// TIA Portal project "ljussennsor skåp" (V18)

(* hardware
DEVICE "S7-1200 station_1"  S7-1200 Station
   slot 0: "Rack_0"  S7-1200 Rack  Rack  V1.0
   slot 1: "PLC_1"  CPU 1212C DC/DC/DC  6ES7 212-1AE40-0XB0  V4.5
DEVICE "HMI_1"  TP900 Comfort
   slot 0: "HMI_1"  TP900 Comfort  6AV2 124-0JC01-0AX0  17.0.0.0
   slot 1: "HMI_RT_1"  TP900 Comfort  6AV2 124-0JC01-0AX0  17.0.0.0
   slot 5: "HMI_1.IE_CP_1"  PROFINET Interface  17.0.0.0
      slot 1: "PROFINET Interface_1"  PROFINET Interface
         slot 1: "Port_1"  Port
         slot 2: "Port_2"  Port
   slot 7: "HMI_1.MPI/DP_CP_1"  MPI/DP Interface  17.0.0.0
*)

// ===== PLC "PLC_1"  CPU 1212C DC/DC/DC =====

VAR_GLOBAL   // PLC tag table "Default tag table"
   "Tag_1" AT %I0.4 : Bool;
   "Tag_2" AT %I0.5 : Bool;
   "Tag_3" AT %I0.6 : Bool;
   "ok" AT %M0.7 : Bool;
END_VAR

VAR_GLOBAL   // PLC tag table "Analog_Tag"
   "Star/Button" AT %I0.0 : Bool;
   "Stop/Button" AT %I0.1 : Bool;
   "Reset/Button" AT %I0.2 : Bool;
   "light sensor" AT %IW64 : Int;
   "Green" AT %Q0.0 : Bool;   // Lamp
   "Red" AT %Q0.1 : Bool;   // Lamp
   "Yellow" AT %Q0.2 : Bool;   // Lamp
   "LEDLights" AT %Q0.3 : Bool;
END_VAR

DATA_BLOCK "data"   // DB1
{ S7_Optimized_Access := 'TRUE' }
VERSION : 0.1
   VAR
      normxstruct : Struct
         minval : Int := 0;
         maxval : Int := 27648;
         lightval : Int;
         normxoutput : Real;
      END_STRUCT;
      lightpercent : Struct
         percentofthelight : Real;
      END_STRUCT;
      calibratedvalues : Struct
         "2layermin" : Real;
         "2layermax" : Real;
      END_STRUCT;
      defaultvalues : Struct
         minimumvalue : Real := 87.9;
         maxvalue : Real := 86.2;
      END_STRUCT;
      startcalibration : Bool;
      finishedcalibration : Bool;
      hmibuttons : Struct
         hmistartbutton : Bool;
         hmiyellowbutton : Bool;
         hmiredbutton : Bool;
      END_STRUCT;
   END_VAR
BEGIN
END_DATA_BLOCK

// folder: System blocks/Program resources

DATA_BLOCK "IEC_Counter_0_DB_1"   // DB3
{ S7_Optimized_Access := 'TRUE' }
AUTHOR : Simatic
FAMILY : IEC
NAME : CNTR
VERSION : 1.0
// stored: InstanceOfName IEC_COUNTER
"IEC_COUNTER"
BEGIN
END_DATA_BLOCK

// folder: (top level)

FUNCTION "function" : Void   // FC1, LAD
{ S7_Optimized_Access := 'TRUE' }
VERSION : 0.1
   VAR_TEMP   // added for the SCL form of the ladder/FBD networks
      _w1 : Bool;
      _w2 : Bool;
      _w3 : Bool;
      _w4 : Bool;
   END_VAR
BEGIN

REGION Network 1: Lamp
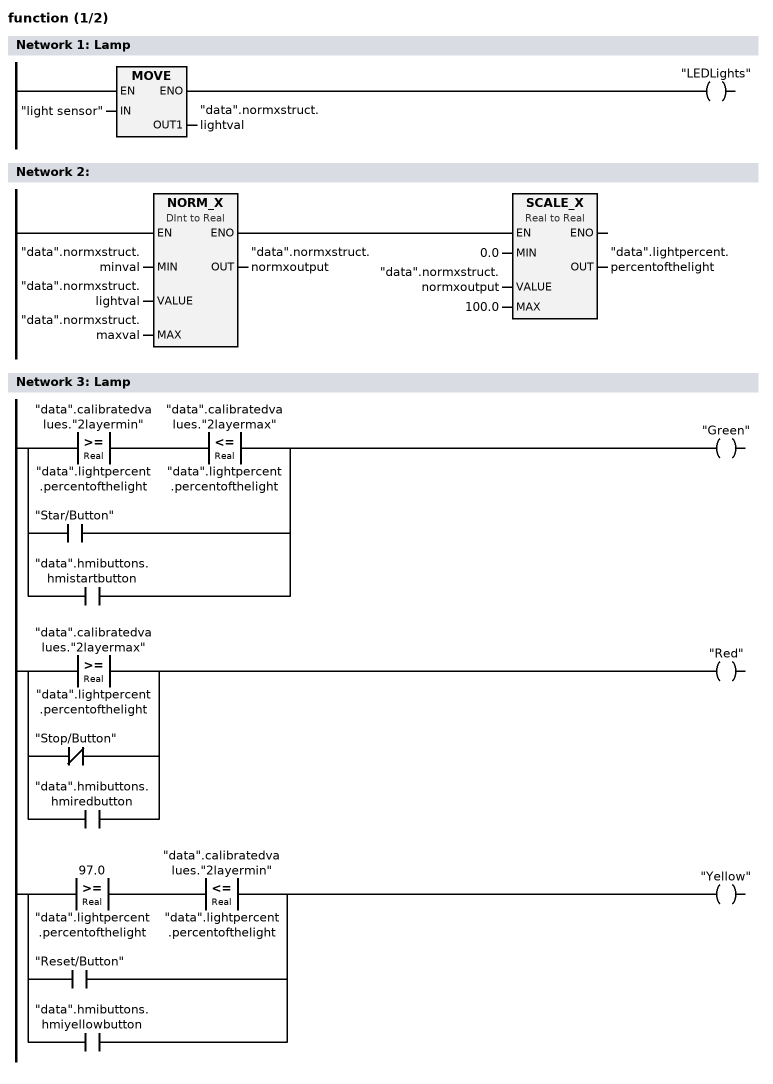
   RUNG wire#powerrail
      Move(in := "light sensor", out1 => "data".normxstruct.lightval)
      Coil( "LEDLights" )
   END_RUNG
   // the same network as SCL:
   "data".normxstruct.lightval := "light sensor";
   "LEDLights" := TRUE;
END_REGION

REGION Network 2
   RUNG wire#powerrail
      { S7_Templates := "[SrcType := DInt, DestType := Real]" } Normalize(min := "data".normxstruct.minval, value := "data".normxstruct.lightval, max := "data".normxstruct.maxval, out => "data".normxstruct.normxoutput)
      { S7_Templates := "[SrcType := Real, DestType := Real]" } Scale(min := 0.0, value := "data".normxstruct.normxoutput, max := 100.0, out => "data".lightpercent.percentofthelight)
   END_RUNG
   // the same network as SCL:
   "data".normxstruct.normxoutput := NORM_X(MIN := "data".normxstruct.minval, VALUE := "data".normxstruct.lightval, MAX := "data".normxstruct.maxval);
   "data".lightpercent.percentofthelight := SCALE_X(MIN := 0.0, VALUE := "data".normxstruct.normxoutput, MAX := 100.0);
END_REGION

REGION Network 3: Lamp
   RUNG wire#powerrail
      { S7_Templates := "SrcType := Real" } GE_Contact(in1 := "data".calibratedvalues."2layermin", in2 := "data".lightpercent.percentofthelight)
      { S7_Templates := "SrcType := Real" } LE_Contact(in1 := "data".calibratedvalues."2layermax", in2 := "data".lightpercent.percentofthelight)
      wire#w1
      Coil( "Green" )
   END_RUNG
   RUNG wire#powerrail
      Contact( "Star/Button" )
   END_RUNG wire#w1
   RUNG wire#powerrail
      Contact( "data".hmibuttons.hmistartbutton )
   END_RUNG wire#w1
   RUNG wire#powerrail
      { S7_Templates := "SrcType := Real" } GE_Contact(in1 := "data".calibratedvalues."2layermax", in2 := "data".lightpercent.percentofthelight)
      wire#w2
      Coil( "Red" )
   END_RUNG
   RUNG wire#powerrail
      I_Contact( "Stop/Button" )
   END_RUNG wire#w2
   RUNG wire#powerrail
      Contact( "data".hmibuttons.hmiredbutton )
   END_RUNG wire#w2
   RUNG wire#powerrail
      { S7_Templates := "SrcType := Real" } GE_Contact(in1 := 97.0, in2 := "data".lightpercent.percentofthelight)
      { S7_Templates := "SrcType := Real" } LE_Contact(in1 := "data".calibratedvalues."2layermin", in2 := "data".lightpercent.percentofthelight)
      wire#w3
      Coil( "Yellow" )
   END_RUNG
   RUNG wire#powerrail
      Contact( "Reset/Button" )
   END_RUNG wire#w3
   RUNG wire#powerrail
      Contact( "data".hmibuttons.hmiyellowbutton )
   END_RUNG wire#w3
   // the same network as SCL:
   "Green" := (("data".calibratedvalues."2layermin" >= "data".lightpercent.percentofthelight) AND ("data".calibratedvalues."2layermax" <= "data".lightpercent.percentofthelight)) OR "Star/Button" OR "data".hmibuttons.hmistartbutton;
   "Red" := ("data".calibratedvalues."2layermax" >= "data".lightpercent.percentofthelight) OR NOT "Stop/Button" OR "data".hmibuttons.hmiredbutton;
   "Yellow" := ((97.0 >= "data".lightpercent.percentofthelight) AND ("data".calibratedvalues."2layermin" <= "data".lightpercent.percentofthelight)) OR "Reset/Button" OR "data".hmibuttons.hmiyellowbutton;
END_REGION

REGION Network 4
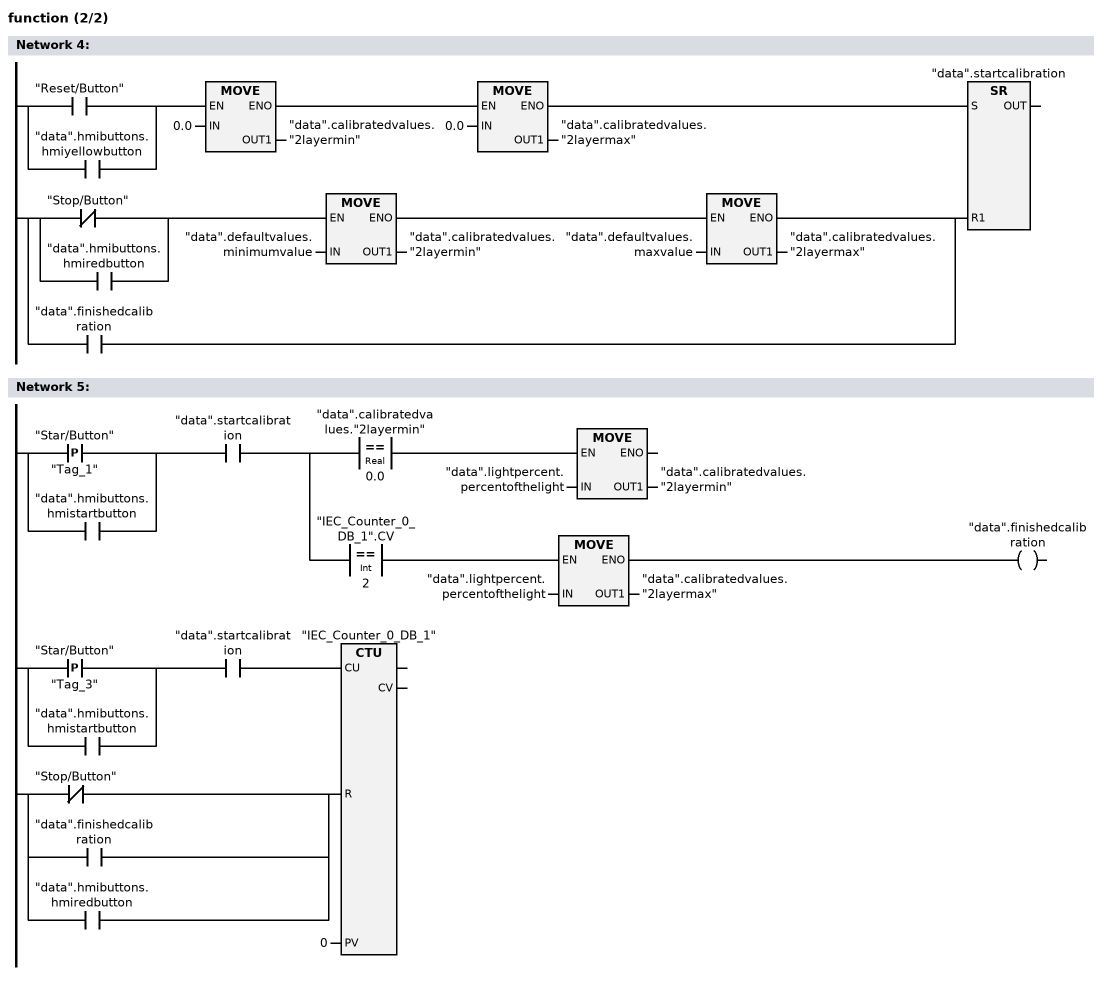
   RUNG wire#powerrail
      Contact( "Reset/Button" )
      wire#w1
      Move(in := 0.0, out1 => "data".calibratedvalues."2layermin")
      Move(in := 0.0, out1 => "data".calibratedvalues."2layermax")
      S_SR(operand := "data".startcalibration, r1 := wire#w3)
   END_RUNG
   RUNG wire#powerrail
      Contact( "data".hmibuttons.hmiyellowbutton )
   END_RUNG wire#w1
   RUNG wire#powerrail
      I_Contact( "Stop/Button" )
      wire#w2
      Move(in := "data".defaultvalues.minimumvalue, out1 => "data".calibratedvalues."2layermin")
      Move(in := "data".defaultvalues.maxvalue, out1 => "data".calibratedvalues."2layermax")
   END_RUNG wire#w3
   RUNG wire#powerrail
      Contact( "data".hmibuttons.hmiredbutton )
   END_RUNG wire#w2
   RUNG wire#powerrail
      Contact( "data".finishedcalibration )
   END_RUNG wire#w3
   // the same network as SCL:
   #_w1 := "Reset/Button" OR "data".hmibuttons.hmiyellowbutton;
   IF #_w1 THEN
       "data".calibratedvalues."2layermin" := 0.0;
       "data".calibratedvalues."2layermax" := 0.0;
   END_IF;
   #_w2 := NOT "Stop/Button" OR "data".hmibuttons.hmiredbutton;
   IF #_w2 THEN
       "data".calibratedvalues."2layermin" := "data".defaultvalues.minimumvalue;
       "data".calibratedvalues."2layermax" := "data".defaultvalues.maxvalue;
   END_IF;
   IF #_w1 THEN
       "data".startcalibration := TRUE;   // SR flip-flop
   END_IF;
   IF #_w2 OR "data".finishedcalibration THEN "data".startcalibration := FALSE; END_IF;
END_REGION

REGION Network 5
   #_w1 := "Star/Button" AND NOT "Tag_1";   // rising edge of "Star/Button"
   "Tag_1" := "Star/Button";
   #_w2 := (#_w1 OR "data".hmibuttons.hmistartbutton) AND "data".startcalibration;
   IF #_w2 AND ("data".calibratedvalues."2layermin" = 0.0) THEN
       "data".calibratedvalues."2layermin" := "data".lightpercent.percentofthelight;
   END_IF;
   #_w3 := #_w2 AND ("IEC_Counter_0_DB_1".CV = 2);
   IF #_w3 THEN "data".calibratedvalues."2layermax" := "data".lightpercent.percentofthelight; END_IF;
   "data".finishedcalibration := #_w3;
   #_w4 := "Star/Button" AND NOT "Tag_3";   // rising edge of "Star/Button"
   "Tag_3" := "Star/Button";
   "IEC_Counter_0_DB_1".CTU(CU := (#_w4 OR "data".hmibuttons.hmistartbutton) AND "data".startcalibration,
                           R := NOT "Stop/Button" OR "data".finishedcalibration OR "data".hmibuttons.hmiredbutton,
                           PV := 0);
END_REGION
END_FUNCTION

ORGANIZATION_BLOCK "Main"   // OB1, LAD, ProgramCycle
TITLE = "Main Program Sweep (Cycle)"
{ S7_Optimized_Access := 'TRUE' }
VERSION : 0.1
   VAR_INPUT
      Initial_Call : Bool;   // Initial call of this OB
      Remanence : Bool;   // =True, if remanent data are available
   END_VAR
BEGIN

REGION Network 1
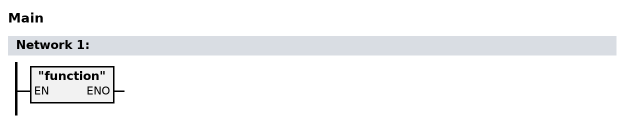
   RUNG wire#powerrail
      "function"()
   END_RUNG
   // the same network as SCL:
   "function"();
END_REGION
END_ORGANIZATION_BLOCK

(* ===== HMI "HMI_RT_1" =====
system functions are stored by id; their names below are inferred from use
connection "Connection_1": ETHERNET, S7_1200_OMS
connection "HMI_Connection_1": ETHERNET, S7_1200_OMS

HMI tags "Default tag table"
   "Tag_ScreenNumber" : UInt, internal
   "Tag_ScreenNumber_1" : UInt, internal
   "greenbuttonhmi" : Bool = PLC data.hmibuttons.hmistartbutton AT %M0.7, 1 s
   "yellowbuttonhmi" : Bool = PLC data.hmibuttons.hmiyellowbutton AT %DB1.DBX0.0, 1 s
   "redbuttonhmi" : Bool = PLC data.hmibuttons.hmiredbutton AT %DB1.DBX0.0, 1 s
   "data_startcalibration" : Bool = PLC data.startcalibration, 1 s

screen "Root screen" 800x420, template "Template_1"
   on GenerateScreen: SetTag("Tag_ScreenNumber", 1)
   Button "Button_1" at 644,23 size 122x64; TextOff 'Calibrate'
      on Press: InvertBit("yellowbuttonhmi")
      on Release: InvertBit("yellowbuttonhmi")
   Button "Button_2" at 644,133 size 122x64; TextOff 'Set'
      on Press: InvertBit("greenbuttonhmi")
      on Release: InvertBit("greenbuttonhmi")
      Appearance <- "data_startcalibration"
   Button "Button_3" at 644,243 size 122x64; TextOff 'Reset'
      on Press: InvertBit("redbuttonhmi")
      on Release: InvertBit("redbuttonhmi")
      Appearance <- "data_startcalibration"

Template "Template_1" 800x420
   Button "Exit" at 720,360 size 78x58; TextOff 'Exit'; PictureOff "ExitRuntime_TP900_Comfort_TR"; PictureOn "ExitRuntime_TP900_Comfort_TR"
      on Release: StopRuntime(0)
   Button "Template_Button" at 640,360 size 78x58; TextOff 'Text'
   Button "Template_Button_1" at 560,360 size 78x58; TextOff 'Text'
   Button "Template_Button_2" at 480,360 size 78x58; TextOff 'Text'
   Button "Template_Button_3" at 400,360 size 78x58; TextOff 'Text'
   Button "Template_Button_4" at 321,360 size 78x58; TextOff 'Text'
   Button "Template_Button_5" at 241,360 size 78x58; TextOff 'Text'
   Button "Template_Button_6" at 161,360 size 78x58; TextOff 'Text'
   Button "Alarms" at 81,360 size 78x58; TextOff 'Alarms'; PictureOff "AlarmDisplay_TP900_Comfort_TR"; PictureOn "AlarmDisplay_TP900_Comfort_TR"
      on Release: function_ef3f5d25("Alarm window_Unacknowledged", -1)
   Button "Start screen" at 1,360 size 78x58; TextOff 'Start screen'; PictureOff "NavigateHome_TP900_Comfort_TR"; PictureOn "NavigateHome_TP900_Comfort_TR"
      on Release: ActivateScreen("Root screen", 0)
*)